// TIA Portal project "Project maybe not work 1.0" (V17) (continued)
REGION Network 7: step 20 Turns on intake and exhaust fans
   "Data_Block_Start_Seq".SeqStep[20] := "Data_Block_Start_Seq".StepNumber = 20;
   "Data_Block_Start_Seq".SeqConditions[20] := ("Data_Block_Start_Seq".StepNumber = 20) AND "FS-115.I" AND "FS-214-I" AND NOT "FS-114.I" AND NOT "FS-213.I" AND "HZ-413.I" AND NOT "PS-411.I" AND NOT "QE-116.I" AND "QE-316.I" AND NOT "Fire lock";
   "Data_Block_Start_Seq".SeqTimer[20].TON(IN := ("Data_Block_Start_Seq".StepNumber = 20) AND "Data_Block_Start_Seq".SeqConditions[20],
                           PT := T#50MS);
   IF "Data_Block_Start_Seq".SeqTimer[20].Q THEN
       "FC" := TRUE;
       "Data_Block_Start_Seq".StepNumber := 25;
   END_IF;
END_REGION

REGION Network 8: step 25 Checks that the fans have turned on
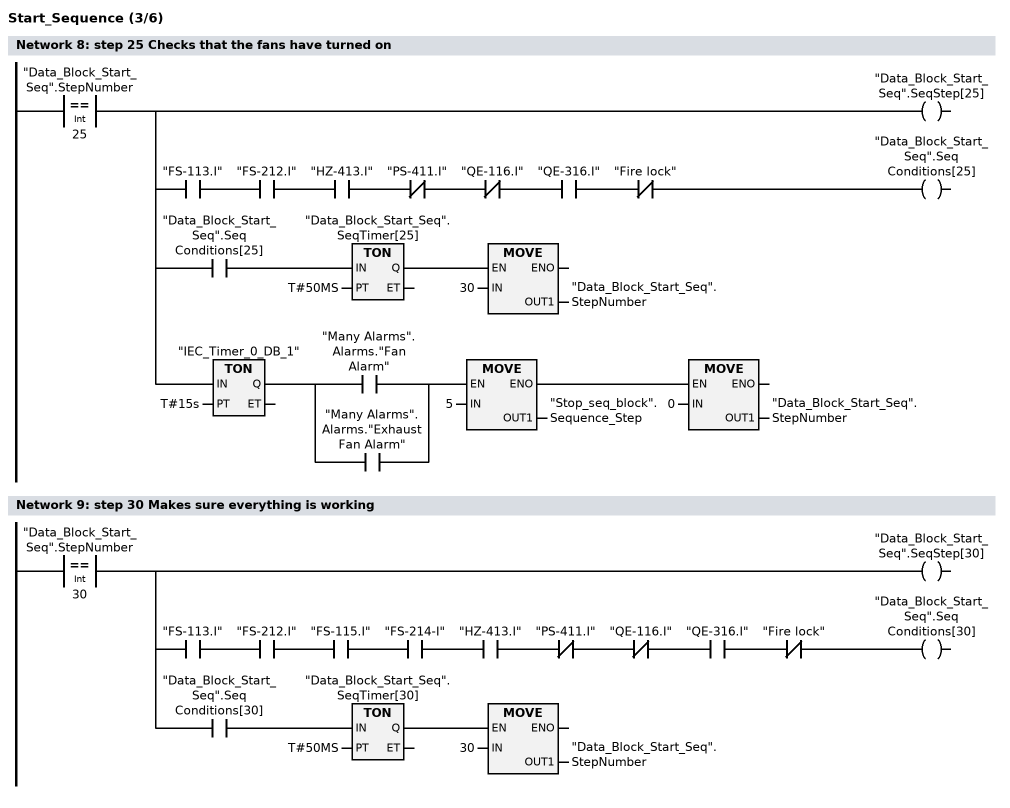
   "Data_Block_Start_Seq".SeqStep[25] := "Data_Block_Start_Seq".StepNumber = 25;
   "Data_Block_Start_Seq".SeqConditions[25] := ("Data_Block_Start_Seq".StepNumber = 25) AND "FS-113.I" AND "FS-212.I" AND "HZ-413.I" AND NOT "PS-411.I" AND NOT "QE-116.I" AND "QE-316.I" AND NOT "Fire lock";
   "Data_Block_Start_Seq".SeqTimer[25].TON(IN := ("Data_Block_Start_Seq".StepNumber = 25) AND "Data_Block_Start_Seq".SeqConditions[25],
                           PT := T#50MS);
   #_w1 := "Data_Block_Start_Seq".StepNumber = 25;
   IF "Data_Block_Start_Seq".SeqTimer[25].Q THEN "Data_Block_Start_Seq".StepNumber := 30; END_IF;
   "IEC_Timer_0_DB_1".TON(IN := #_w1, PT := T#15s);
   IF "IEC_Timer_0_DB_1".Q AND ("Many Alarms".Alarms."Fan Alarm" OR "Many Alarms".Alarms."Exhaust Fan Alarm") THEN
       "Stop_seq_block".Sequence_Step := 5;
       "Data_Block_Start_Seq".StepNumber := 0;
   END_IF;
END_REGION

REGION Network 9: step 30 Makes sure everything is working
   "Data_Block_Start_Seq".SeqStep[30] := "Data_Block_Start_Seq".StepNumber = 30;
   "Data_Block_Start_Seq".SeqConditions[30] := ("Data_Block_Start_Seq".StepNumber = 30) AND "FS-113.I" AND "FS-212.I" AND "FS-115.I" AND "FS-214-I" AND "HZ-413.I" AND NOT "PS-411.I" AND NOT "QE-116.I" AND "QE-316.I" AND NOT "Fire lock";
   "Data_Block_Start_Seq".SeqTimer[30].TON(IN := ("Data_Block_Start_Seq".StepNumber = 30) AND "Data_Block_Start_Seq".SeqConditions[30],
                           PT := T#50MS);
   IF "Data_Block_Start_Seq".SeqTimer[30].Q THEN "Data_Block_Start_Seq".StepNumber := 30; END_IF;
END_REGION

REGION Network 10: step 30 Makes sure everything is working
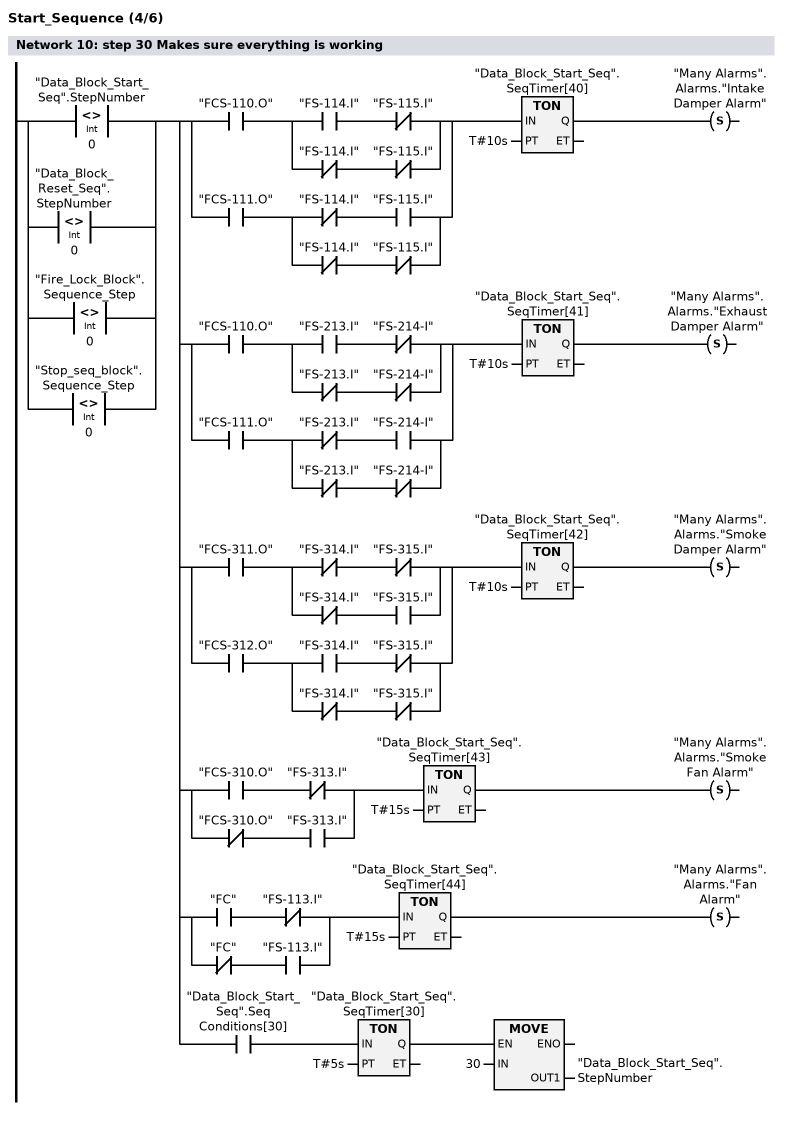
   #_w1 := ("Data_Block_Start_Seq".StepNumber <> 0) OR ("Data_Block_Reset_Seq".StepNumber <> 0) OR ("Fire_Lock_Block".Sequence_Step <> 0) OR ("Stop_seq_block".Sequence_Step <> 0);
   "Data_Block_Start_Seq".SeqTimer[40].TON(IN := #_w1 AND (("FCS-110.O" AND (("FS-114.I" AND NOT "FS-115.I") OR (NOT "FS-114.I" AND NOT "FS-115.I"))) OR ("FCS-111.O" AND ((NOT "FS-114.I" AND "FS-115.I") OR (NOT "FS-114.I" AND NOT "FS-115.I")))),
                           PT := T#10s);
   IF "Data_Block_Start_Seq".SeqTimer[40].Q THEN "Many Alarms".Alarms."Intake Damper Alarm" := TRUE; END_IF;
   "Data_Block_Start_Seq".SeqTimer[41].TON(IN := #_w1 AND (("FCS-110.O" AND (("FS-213.I" AND NOT "FS-214-I") OR (NOT "FS-213.I" AND NOT "FS-214-I"))) OR ("FCS-111.O" AND ((NOT "FS-213.I" AND "FS-214-I") OR (NOT "FS-213.I" AND NOT "FS-214-I")))),
                           PT := T#10s);
   IF "Data_Block_Start_Seq".SeqTimer[41].Q THEN "Many Alarms".Alarms."Exhaust Damper Alarm" := TRUE; END_IF;
   "Data_Block_Start_Seq".SeqTimer[42].TON(IN := #_w1 AND (("FCS-311.O" AND ((NOT "FS-314.I" AND NOT "FS-315.I") OR (NOT "FS-314.I" AND "FS-315.I"))) OR ("FCS-312.O" AND (("FS-314.I" AND NOT "FS-315.I") OR (NOT "FS-314.I" AND NOT "FS-315.I")))),
                           PT := T#10s);
   IF "Data_Block_Start_Seq".SeqTimer[42].Q THEN "Many Alarms".Alarms."Smoke Damper Alarm" := TRUE; END_IF;
   "Data_Block_Start_Seq".SeqTimer[43].TON(IN := #_w1 AND (("FCS-310.O" AND NOT "FS-313.I") OR (NOT "FCS-310.O" AND "FS-313.I")),
                           PT := T#15s);
   IF "Data_Block_Start_Seq".SeqTimer[43].Q THEN "Many Alarms".Alarms."Smoke Fan Alarm" := TRUE; END_IF;
   "Data_Block_Start_Seq".SeqTimer[44].TON(IN := #_w1 AND (("FC" AND NOT "FS-113.I") OR (NOT "FC" AND "FS-113.I")),
                           PT := T#15s);
   IF "Data_Block_Start_Seq".SeqTimer[44].Q THEN "Many Alarms".Alarms."Fan Alarm" := TRUE; END_IF;
   "Data_Block_Start_Seq".SeqTimer[30].TON(IN := #_w1 AND "Data_Block_Start_Seq".SeqConditions[30], PT := T#5s);
   IF "Data_Block_Start_Seq".SeqTimer[30].Q THEN "Data_Block_Start_Seq".StepNumber := 30; END_IF;
END_REGION

REGION Network 11: Stop and reset button function. after 3s puts on stop sequence if 10s passes reset function turns on
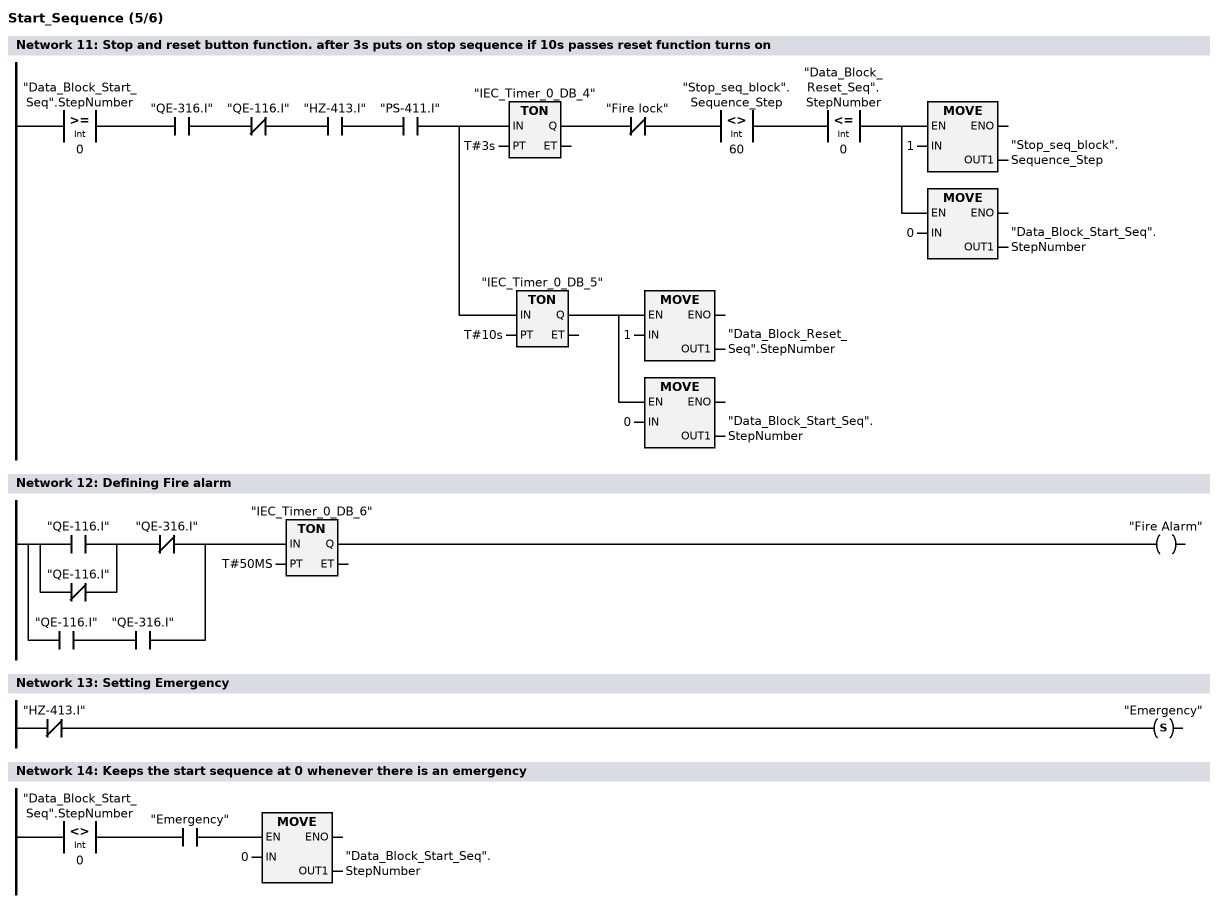
   #_w1 := ("Data_Block_Start_Seq".StepNumber >= 0) AND "QE-316.I" AND NOT "QE-116.I" AND "HZ-413.I" AND "PS-411.I";
   "IEC_Timer_0_DB_4".TON(IN := #_w1, PT := T#3s);
   #_w2 := "IEC_Timer_0_DB_4".Q AND NOT "Fire lock" AND ("Stop_seq_block".Sequence_Step <> 60) AND ("Data_Block_Reset_Seq".StepNumber <= 0);
   IF #_w2 THEN
       "Stop_seq_block".Sequence_Step := 1;
       "Data_Block_Start_Seq".StepNumber := 0;
   END_IF;
   "IEC_Timer_0_DB_5".TON(IN := #_w1, PT := T#10s);
   IF "IEC_Timer_0_DB_5".Q THEN
       "Data_Block_Reset_Seq".StepNumber := 1;
       "Data_Block_Start_Seq".StepNumber := 0;
   END_IF;
END_REGION

REGION Network 12: Defining Fire alarm
   "IEC_Timer_0_DB_6".TON(IN := (("QE-116.I" OR NOT "QE-116.I") AND NOT "QE-316.I") OR ("QE-116.I" AND "QE-316.I"),
                          PT := T#50MS);
   "Fire Alarm" := "IEC_Timer_0_DB_6".Q;
END_REGION

REGION Network 13: Setting Emergency
   RUNG wire#powerrail
      I_Contact( "HZ-413.I" )
      S_Coil( "Emergency" )
   END_RUNG
   // the same network as SCL:
   IF NOT "HZ-413.I" THEN "Emergency" := TRUE; END_IF;
END_REGION

REGION Network 14: Keeps the start sequence at 0 whenever there is an emergency
   RUNG wire#powerrail
      { S7_Templates := "SrcType := Int" } NE_Contact(in1 := "Data_Block_Start_Seq".StepNumber, in2 := 0)
      Contact( "Emergency" )
      Move(in := 0, out1 => "Data_Block_Start_Seq".StepNumber)
   END_RUNG
   // the same network as SCL:
   IF ("Data_Block_Start_Seq".StepNumber <> 0) AND "Emergency" THEN
       "Data_Block_Start_Seq".StepNumber := 0;
   END_IF;
END_REGION

REGION Network 15: Defining Alarm
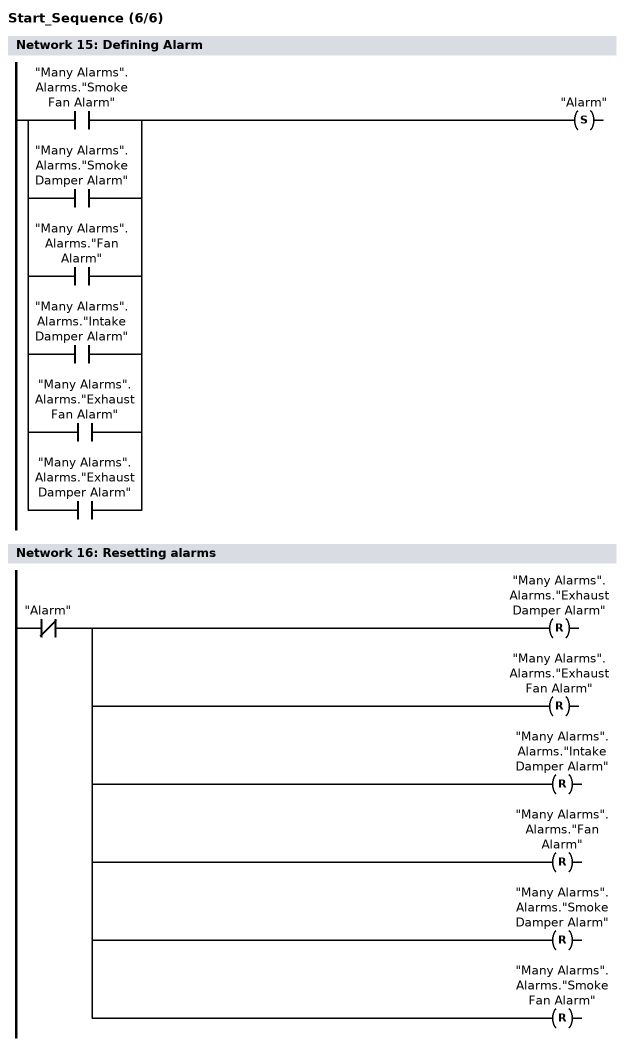
   RUNG wire#powerrail
      Contact( "Many Alarms".Alarms."Smoke Fan Alarm" )
      wire#w1
      S_Coil( "Alarm" )
   END_RUNG
   RUNG wire#powerrail
      Contact( "Many Alarms".Alarms."Smoke Damper Alarm" )
   END_RUNG wire#w1
   RUNG wire#powerrail
      Contact( "Many Alarms".Alarms."Fan Alarm" )
   END_RUNG wire#w1
   RUNG wire#powerrail
      Contact( "Many Alarms".Alarms."Intake Damper Alarm" )
   END_RUNG wire#w1
   RUNG wire#powerrail
      Contact( "Many Alarms".Alarms."Exhaust Fan Alarm" )
   END_RUNG wire#w1
   RUNG wire#powerrail
      Contact( "Many Alarms".Alarms."Exhaust Damper Alarm" )
   END_RUNG wire#w1
   // the same network as SCL:
   IF "Many Alarms".Alarms."Smoke Fan Alarm" OR "Many Alarms".Alarms."Smoke Damper Alarm" OR "Many Alarms".Alarms."Fan Alarm" OR "Many Alarms".Alarms."Intake Damper Alarm" OR "Many Alarms".Alarms."Exhaust Fan Alarm" OR "Many Alarms".Alarms."Exhaust Damper Alarm" THEN
       "Alarm" := TRUE;
   END_IF;
END_REGION

REGION Network 16: Resetting alarms
   RUNG wire#powerrail
      I_Contact( "Alarm" )
      wire#w1
      R_Coil( "Many Alarms".Alarms."Exhaust Damper Alarm" )
   END_RUNG
   RUNG wire#w1
      R_Coil( "Many Alarms".Alarms."Exhaust Fan Alarm" )
   END_RUNG
   RUNG wire#w1
      R_Coil( "Many Alarms".Alarms."Intake Damper Alarm" )
   END_RUNG
   RUNG wire#w1
      R_Coil( "Many Alarms".Alarms."Fan Alarm" )
   END_RUNG
   RUNG wire#w1
      R_Coil( "Many Alarms".Alarms."Smoke Damper Alarm" )
   END_RUNG
   RUNG wire#w1
      R_Coil( "Many Alarms".Alarms."Smoke Fan Alarm" )
   END_RUNG
   // the same network as SCL:
   IF NOT "Alarm" THEN
       "Many Alarms".Alarms."Exhaust Damper Alarm" := FALSE;
       "Many Alarms".Alarms."Exhaust Fan Alarm" := FALSE;
       "Many Alarms".Alarms."Intake Damper Alarm" := FALSE;
       "Many Alarms".Alarms."Fan Alarm" := FALSE;
       "Many Alarms".Alarms."Smoke Damper Alarm" := FALSE;
       "Many Alarms".Alarms."Smoke Fan Alarm" := FALSE;
   END_IF;
END_REGION
END_FUNCTION

ORGANIZATION_BLOCK "Main"   // OB1, LAD, ProgramCycle
TITLE = "Main Program Sweep (Cycle)"
{ S7_Optimized_Access := 'TRUE' }
VERSION : 0.1
   VAR_INPUT
      Initial_Call : Bool;   // Initial call of this OB
      Remanence : Bool;   // =True, if remanent data are available
   END_VAR
   VAR_TEMP
      "QE.200i-norm" : Real;
   END_VAR
   VAR_TEMP   // added for the SCL form of the ladder/FBD networks
      _w1 : Bool;
      _w2 : Bool;
      _w3 : Bool;
   END_VAR
BEGIN

REGION Network 1
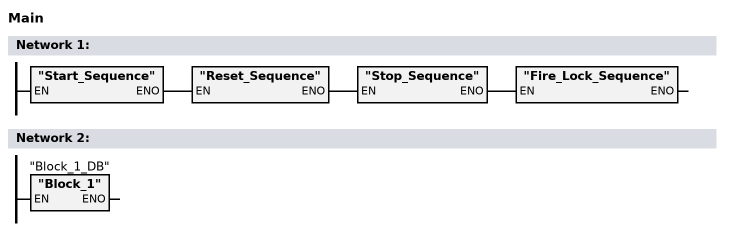
   RUNG wire#powerrail
      "Start_Sequence"()
      "Reset_Sequence"()
      "Stop_Sequence"()
      "Fire_Lock_Sequence"()
   END_RUNG
   // the same network as SCL:
   "Start_Sequence"(ENO => #_w1);
   "Reset_Sequence"(EN := #_w1, ENO => #_w2);
   "Stop_Sequence"(EN := #_w2, ENO => #_w3);
   IF #_w3 THEN "Fire_Lock_Sequence"(); END_IF;
END_REGION

REGION Network 2
   RUNG wire#powerrail
      "Block_1_DB"()
   END_RUNG
   // the same network as SCL:
   "Block_1_DB"();   // "Block_1"
END_REGION
END_ORGANIZATION_BLOCK

ORGANIZATION_BLOCK "Cyclic interrupt"   // OB30, LAD, CyclicInterrupt
{ S7_Optimized_Access := 'TRUE' }
VERSION : 0.1
   VAR_INPUT
      Initial_Call : Bool;   // Initial call of this OB
      Event_Count : Int;   // Events discarded
   END_VAR
   VAR_TEMP
      QE_Temp : Real;
      "TE temp" : Real;
      "TFC-Output temp" : Real;
   END_VAR
BEGIN

REGION Network 1
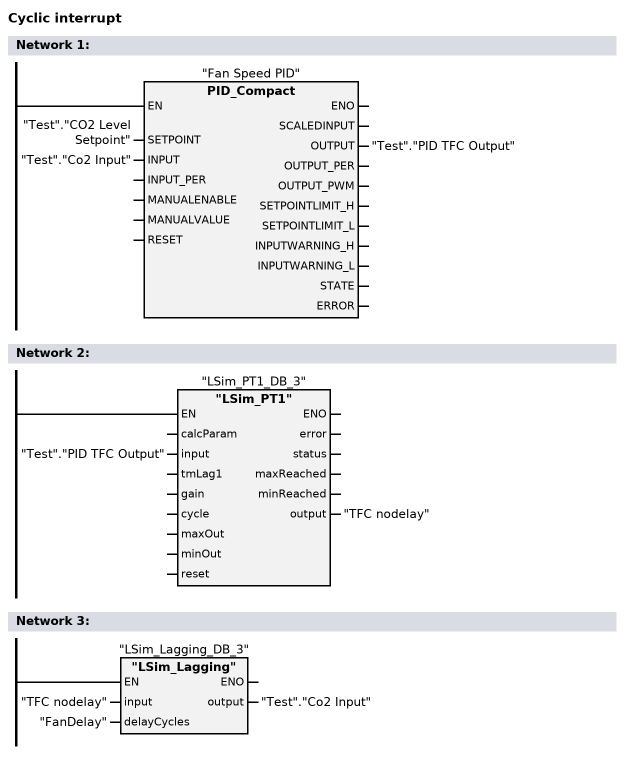
   "Fan Speed PID"(Setpoint := "Test"."CO2 Level Setpoint",   // PID_Compact
                   Input := "Test"."Co2 Input",
                   Output => "Test"."PID TFC Output");
END_REGION

REGION Network 2
   RUNG wire#powerrail
      "LSim_PT1_DB_3"(calcParam :=, input := "Test"."PID TFC Output", tmLag1 :=, gain :=, cycle :=, maxOut :=, minOut :=, reset :=, error =>, status =>, maxReached =>, minReached =>, output => "TFC nodelay")
   END_RUNG
   // the same network as SCL:
   "LSim_PT1_DB_3"(input := "Test"."PID TFC Output", output => "TFC nodelay");   // "LSim_PT1"
END_REGION

REGION Network 3
   RUNG wire#powerrail
      "LSim_Lagging_DB_3"(input := "TFC nodelay", delayCycles := "FanDelay", output => "Test"."Co2 Input")
   END_RUNG
   // the same network as SCL:
   "LSim_Lagging_DB_3"(input := "TFC nodelay", delayCycles := "FanDelay", output => "Test"."Co2 Input");   // "LSim_Lagging"
END_REGION
END_ORGANIZATION_BLOCK

ORGANIZATION_BLOCK "Cyclic interrupt_1"   // OB31, LAD, CyclicInterrupt
{ S7_Optimized_Access := 'TRUE' }
VERSION : 0.1
   VAR_INPUT
      Initial_Call : Bool;   // Initial call of this OB
      Event_Count : Int;   // Events discarded
   END_VAR
BEGIN

REGION Network 1
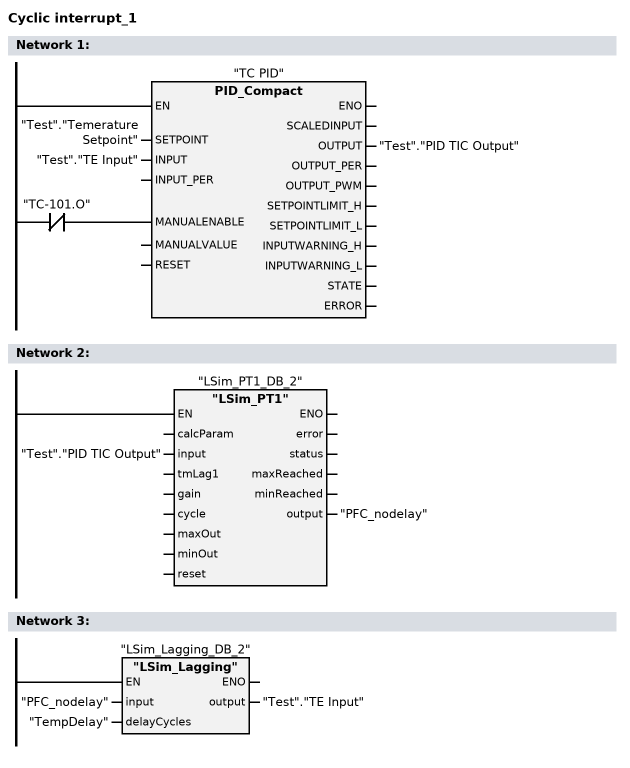
   "TC PID"(Setpoint := "Test"."Temerature Setpoint",   // PID_Compact
            Input := "Test"."TE Input",
            ManualEnable := NOT "TC-101.O",
            Output => "Test"."PID TIC Output");
END_REGION

REGION Network 2
   RUNG wire#powerrail
      "LSim_PT1_DB_2"(calcParam :=, input := "Test"."PID TIC Output", tmLag1 :=, gain :=, cycle :=, maxOut :=, minOut :=, reset :=, error =>, status =>, maxReached =>, minReached =>, output => "PFC_nodelay")
   END_RUNG
   // the same network as SCL:
   "LSim_PT1_DB_2"(input := "Test"."PID TIC Output", output => "PFC_nodelay");   // "LSim_PT1"
END_REGION

REGION Network 3
   RUNG wire#powerrail
      "LSim_Lagging_DB_2"(input := "PFC_nodelay", delayCycles := "TempDelay", output => "Test"."TE Input")
   END_RUNG
   // the same network as SCL:
   "LSim_Lagging_DB_2"(input := "PFC_nodelay", delayCycles := "TempDelay", output => "Test"."TE Input");   // "LSim_Lagging"
END_REGION
END_ORGANIZATION_BLOCK

(* ===== HMI "HMI_RT_1" =====
system functions are stored by id; their names below are inferred from use
connection "HMI_Connection_1": ETHERNET, S7_1200_OMS
connection "HMI_Connection_2": ETHERNET, S7_1200_OMS

HMI tags "Default tag table"
   "Tag_ScreenNumber" : UInt, internal
   "Fire lock" : Bool = PLC "Fire lock" AT %M36.2, 1 s
   "Emergency" : Bool = PLC Emergency AT %M36.4, 1 s
   "Intake Fan" : Bool = PLC "FS-113.I" AT %I6.1, 1 s
   "Exhaust Fan" : Bool = PLC "FS-212.I" AT %I6.4, 1 s
   "Intake Damper Closing" : Bool = PLC "FCS-111.O" AT %Q0.2, 1 s
   "Intake Damper Opening" : Bool = PLC "FCS-110.O" AT %Q0.1, 1 s
   "Intake Damper Closed" : Bool = PLC "FS-114.I" AT %I7.5, 1 s
   "Intake Damper Open" : Bool = PLC "FS-115.I" AT %I7.1, 1 s
   "Exhaust Damper Closing" : Bool = PLC "FCS-211.O" AT %Q0.4, 1 s
   "Exhaust Damper Closed" : Bool = PLC "FS-213.I" AT %I7.4, 1 s
   "Exhaust Damper Opening" : Bool = PLC "FCS-210O" AT %Q0.3, 1 s
   "Exhaust Damper Open" : Bool = PLC "FS-214-I" AT %I7.0, 1 s
   "Smoke Damper Opening" : Bool = PLC "FCS-311.O" AT %Q0.6, 1 s
   "Smoke Damper Open" : Bool = PLC "FS-314.I" AT %I7.2, 1 s
   "Smoke Damper Closing" : Bool = PLC "FCS-312.O" AT %Q0.7, 1 s
   "Smoke Damper Closed" : Bool = PLC "FS-315.I" AT %I7.6, 1 s
   "Smoke Fan Control" : Bool = PLC "FCS-310.O" AT %Q0.5, 1 s
   "Start Button" : Bool = PLC "PS-410.I" AT %I6.0, 1 s
   "Stop/Reset Button" : Bool = PLC "PS-411.I" AT %I6.3, 1 s
   "Emergency Button" : Bool = PLC "HZ-413.I" AT %I6.5, 1 s
   "Start Seq" : Int = PLC Data_Block_Start_Seq.StepNumber AT %DB1.DBX0.0, 1 s
   "Stop Seq" : Int = PLC Stop_seq_block.Sequence_Step AT %DB1.DBX0.0, 1 s
   "Reset Seq" : Int = PLC Data_Block_Reset_Seq.StepNumber AT %DB1.DBX0.0, 1 s
   "Fire Lock Seq" : Int = PLC Fire_Lock_Block.Sequence_Step AT %M36.2, 1 s
   "Fire Inside" : Bool = PLC "QE-316.I" AT %I7.7, 1 s
   "Fire Outside" : Bool = PLC "QE-116.I" AT %I7.3, 1 s
   "Smoke Fan Status" : Bool = PLC "FS-313.I" AT %I6.2, 1 s
   "Intake Fan Control" : Bool = PLC FC AT %M20.0, 1 s
   "Speed Scale" : Int = PLC Test."CO2 Level Setpoint" AT %DB1.DBW0, 1 s
   "TFC-201sp" : Real = PLC "Co2 Setpoint" AT %MD200, 1 s
   "QE-200.i" : Int = PLC "QE-200.i" AT %MW64, 1 s
   "TFC-201.o" : Real = PLC "TFC-201.o" AT %MD80, 1 s
   "Temperature.sp" : Int = PLC "Temperature.sp" AT %MW222, 1 s
   "TE-100.i" : Int = PLC "TE-100.i" AT %MW66, 1 s
   "TempratureSp" : Int = PLC "Temperature.sp" AT %MW222, 1 s
   "PFC-202.o" : Real = PLC "PFC-202.o" AT %MD84, 1 s
   "Test_PID_Data_Output" : Real = PLC Test."PID TFC Output", 1 s
   "Fan Speed PID_Output" : Real = PLC "Fan Speed PID".Output, 1 s
   "Fan Speed PID_Input" : Real = PLC "Fan Speed PID".Input, 1 s
   "Data_Block_Start_Seq_SeqStep{5}" : Bool = PLC Data_Block_Start_Seq.SeqStep[5], 1 s
   "Test_Temerature Setpoint" : Int = PLC Test."Temerature Setpoint", 1 s
   "TC PID_Input" : Real = PLC "TC PID".Input, 1 s
   "Fan Speed PID_State" : Int = PLC "Fan Speed PID".State, 1 s
   "TC PID_State" : Int = PLC "TC PID".State, 1 s

HMI tags "Alarms"
   "Alarms" : Int AT %DB4.DBW0, 1 s

discrete alarms
   1: 'Wha', class Warnings, trigger "Alarms" bit 0
   2: 'Wha', class Warnings, trigger "Alarms" bit 1
   3: 'Wha', class Warnings, trigger "Alarms" bit 2
   4: 'Wha', class Warnings, trigger "Alarms" bit 3
   5: 'Wha', class Warnings, trigger "Alarms" bit 4
   6: 'Wha', class Warnings, trigger "Alarms" bit 5
   7: 'Wha', class Warnings, trigger "Alarms" bit 6
   8: 'Wha', class Warnings, trigger "Alarms" bit 7
   9: 'Intake Damper Control Time Exceeded', class Errors, trigger "Alarms" bit 8
   10: 'Intake Fan Control Time Exceeded', class Errors, trigger "Alarms" bit 9
   13: 't Dameper Control Time Exceeded', class Errors, trigger "Alarms" bit 10
   14: 'Exhaust Fan Control time Exceeded', class Errors, trigger "Alarms" bit 11
   15: 'Smoke Damper Control Time Exceeded', class Errors, trigger "Alarms" bit 12
   16: 'Smoke Fan Control Time Exceeded', class Errors, trigger "Alarms" bit 13

screen "Root screen" 1280x757, template "Template_1"
   on GenerateScreen: SetTag("Tag_ScreenNumber", 1)
   Circle "Circle_1" at 336,50 size 29x29
      Appearance <- "Fire lock"
   Circle "Circle_2" at 334,83 size 29x29
      Appearance <- "Emergency"
      Visibility <- "Emergency"
   Button "HmiScreenItemData_2" at 36,95 size 159x47; TextOff 'System screens'; PictureOff "Navigates to System screens for TP2200 Comfort V2 17.0.0.0"; PictureOn "Navigates to System screens for TP2200 Comfort V2 17.0.0.0"
      on Release: ActivateScreen("System screens", 0)
   Button "HmiScreenItemData" at 36,36 size 159x47; TextOff 'Screen0'; PictureOff "Navigates to Screen0 for TP2200 Comfort V2 17.0.0.0"; PictureOn "Navigates to Screen0 for TP2200 Comfort V2 17.0.0.0"
      on Release: ActivateScreen("Screen0", 0)
   Rectangle "Exhaust Damper Opening" at 833,244 size 54x23
      Appearance <- "Exhaust Damper Opening"
      Visibility <- "Exhaust Damper Opening"
   Rectangle "Intake Damper Opening" at 542,400 size 54x23
      Appearance <- "Intake Damper Opening"
      Visibility <- "Intake Damper Opening"
   Rectangle "Intake Damper Closing" at 542,400 size 54x23
      Appearance <- "Intake Damper Closing"
      Visibility <- "Intake Damper Closing"
   Rectangle "Exhaust Damper Closing" at 833,244 size 54x23
      Appearance <- "Exhaust Damper Closing"
      Visibility <- "Exhaust Damper Closing"
   Circle "Circle_3" at 334,83 size 29x29
      Appearance <- "Emergency Button"
      Visibility <- "Emergency Button"
   Rectangle "Smoke Damper Closing" at 833,149 size 54x23
      Appearance <- "Smoke Damper Closing"
      Visibility <- "Smoke Damper Closing"
   Rectangle "Smoke Damper Opening" at 833,149 size 54x23
      Appearance <- "Smoke Damper Opening"
      Visibility <- "Smoke Damper Opening"
   Button "Smoke Damper Closed Button_1" at 210,565 size 96x32; TextOff 'Closed'
      on Click: SetBit("Smoke Damper Closed")
      Visibility <- "Smoke Damper Closed"
   Button "Smoke Damper Open Button_1" at 210,610 size 96x32; TextOff 'Open'
      on Click: SetBit("Smoke Damper Open")
      Visibility <- "Smoke Damper Open"
   Button "Smoke Damper Not Closed Button_1" at 210,566 size 96x32; TextOff 'Not Closed'
      on Click: ResetBit("Smoke Damper Closed")
      Visibility <- "Smoke Damper Closed"
   Button "Smoke Damper Not Open Button_1" at 210,609 size 96x32; TextOff 'Not Open'
      on Click: ResetBit("Smoke Damper Open")
      Visibility <- "Smoke Damper Open"
   Button "Intake Damper Closed Button" at 7,565 size 96x32; TextOff 'Closed'
      on Click: SetBit("Intake Damper Closed")
      Visibility <- "Intake Damper Closed"
   Button "Intake Damper Open Button" at 7,610 size 96x32; TextOff 'Open'
      on Click: SetBit("Intake Damper Open")
      Visibility <- "Intake Damper Open"
   Button "Intake Damper Not Closed Button" at 8,565 size 96x32; TextOff 'Not Closed'
      on Click: ResetBit("Intake Damper Closed")
      Visibility <- "Intake Damper Closed"
   Button "Exhaust Damper Closed Button" at 108,565 size 96x32; TextOff 'Closed'
      on Click: SetBit("Exhaust Damper Closed")
      Visibility <- "Exhaust Damper Closed"
   Button "Intake Damper Not Open Button" at 7,608 size 96x32; TextOff 'Not Open'
      Visibility <- "Intake Damper Open"
      on Click: ResetBit("Intake Damper Open")
   Button "Exhaust Damper Open Button" at 108,610 size 96x32; TextOff 'Open'
      on Click: SetBit("Exhaust Damper Open")
      Visibility <- "Exhaust Damper Open"
   Button "Exhaust Damper Not Closed Button" at 108,565 size 96x32; TextOff 'Not Closed'
      on Click: ResetBit("Exhaust Damper Closed")
      Visibility <- "Exhaust Damper Closed"
   Button "Exhaust Damper Not Open Button" at 108,608 size 96x32; TextOff 'Not Open'
      on Click: ResetBit("Exhaust Damper Open")
      Visibility <- "Exhaust Damper Open"
   GraphicView "Graphic view_1" at 430,120 size 824x564; Picture "Graphic_10"
   Rectangle "Exhaust Fan" at 650,229 size 54x23
      Appearance <- "Intake Fan Control"
   Rectangle "Intake Fan" at 730,383 size 54x23
      Appearance <- "Intake Fan Control"
   Rectangle "Intake Damper Closed" at 542,400 size 54x23
      Appearance <- "Intake Damper Closed"
      Visibility <- "Intake Damper Closed"
   Rectangle "Intake Damper Open" at 542,400 size 54x23
      Appearance <- "Intake Damper Open"
      Visibility <- "Intake Damper Open"
   Rectangle "Exhaust Damper Open" at 833,244 size 54x23
      Appearance <- "Exhaust Damper Open"
      Visibility <- "Exhaust Damper Open"
   Rectangle "Exhaust Damper Closed" at 833,244 size 54x23
      Visibility <- "Exhaust Damper Closed"
      Appearance <- "Exhaust Damper Closed"
   Rectangle "Smoke Damper Open" at 833,149 size 54x23
      Appearance <- "Smoke Damper Open"
      Visibility <- "Smoke Damper Open"
   Rectangle "Smoke Damper Closed" at 833,149 size 54x23
      Visibility <- "Smoke Damper Closed"
      Appearance <- "Smoke Damper Closed"
   Button "Intake Fan Off" at 7,648 size 96x32; TextOff 'OFF'
      on Click: ResetBit("Intake Fan")
      Visibility <- "Intake Fan"
   Button "Intake Fan On" at 7,648 size 96x32; TextOff 'ON'
      on Click: SetBit("Intake Fan")
      Visibility <- "Intake Fan"
   Button "Exhaust Fan Off" at 108,648 size 96x32; TextOff 'OFF'
      on Click: ResetBit("Exhaust Fan")
      Visibility <- "Exhaust Fan"
   Button "Exhaust Fan on" at 108,648 size 96x32; TextOff 'ON'
      on Click: SetBit("Exhaust Fan")
      Visibility <- "Exhaust Fan"
   Button "Button_1" at 47,162 size 210x95; TextOff 'Start'
      on Press: SetBit("Start Button")
      on Release: ResetBit("Start Button")
      Appearance <- "Data_Block_Start_Seq_SeqStep{5}"
   Button "Button_2" at 47,272 size 210x45; TextOff 'Stop/Reset'
      on Press: SetBit("Stop/Reset Button")
      on Release: ResetBit("Stop/Reset Button")
   Button "Button_3" at 45,340 size 210x45; TextOff 'Release Emergency'
      on Click: SetBit("Emergency Button")
   Button "Button_4" at 45,387 size 210x45; TextOff 'Emergency'
      on Click: ResetBit("Emergency Button")
   Rectangle "Rectangle_1" at 416,67 size 50x45
      Appearance <- "Start Seq"
   Rectangle "Rectangle_2" at 479,65 size 50x45
      Appearance <- "Stop Seq"
   Rectangle "Rectangle_3" at 544,67 size 50x45
      Appearance <- "Reset Seq"
   Rectangle "Rectangle_4" at 607,65 size 50x45
      Appearance <- "Fire Lock Seq"
   Button "Button_5" at 35,480 size 96x32; TextOff 'Fire O'
      on Click: SetBit("Fire Outside")
      Visibility <- "Fire Outside"
   Button "Button_6" at 32,480 size 96x32; TextOff 'No Fire O'
      on Click: ResetBit("Fire Outside")
      Visibility <- "Fire Outside"
   Button "Button_7" at 177,480 size 96x32; TextOff 'Fire I'
      on Click: ResetBit("Fire Inside")
      Visibility <- "Fire Inside"
   Button "Button_8" at 178,480 size 96x32; TextOff 'No Fire I'
      on Click: SetBit("Fire Inside")
      Visibility <- "Fire Inside"
   Rectangle "Rectangle_5" at 35,443 size 95x24
      Appearance <- "Fire Outside"
   Rectangle "Rectangle_6" at 180,442 size 95x24
      Appearance <- "Fire Inside"
   Rectangle "Smoke Exhaust Fan_1" at 652,133 size 54x23
      Appearance <- "Smoke Fan Control"
   TextField "Text field_1" at 23,540 size 67x25; Text 'Intake'
   TextField "Text field_2" at 115,540 size 80x25; Text 'Exhaust'
   TextField "Text field_3" at 225,540 size 68x25; Text 'Smoke'
   Button "Smoke Fan Off" at 210,648 size 96x32; TextOff 'OFF'
      on Click: ResetBit("Smoke Fan Status")
      Visibility <- "Smoke Fan Status"
   Button "Smoke Fan On" at 210,648 size 96x32; TextOff 'ON'
      on Click: SetBit("Smoke Fan Status")
      Visibility <- "Smoke Fan Status"
   Button "Button_10" at 649,256 size 64x61; TextOff 'Text'; TextOn 'Exhaust Fan Speed'
      on Click: function_efd93a16("Fan Speed", 0, 0, -1, -1, 1)
   Button "Button_11" at 890,402 size 151x79; TextOff 'Text'; TextOn 'Pop-up screen_1'
      on Click: function_efd93a16("Pop-up screen_1", 0, 0, -1, -1, 1)
   Bar "Bar_1" at 1147,164 size 80x230; MinimumValue 0; MaximumValue 100
      ProcessValue <- "Fan Speed PID_Input"
   IOField "I/O field_1" at 1142,405 size 96x32; FormatPattern 999; Unit %
      ProcessValue <- "Speed Scale"
   TextField "Text field_4" at 1162,138 size 43x25; Text 'CO2'
   Button "Button_9" at 733,412 size 55x58; TextOn 'Exhaust Fan Speed'; TextOff 'Text'
      on Click: function_efd93a16("Fan Speed", 0, 0, -1, -1, 1)
   IOField "I/O field_2" at 1142,459 size 96x32; FormatPattern s99999
      ProcessValue <- "Fan Speed PID_State"
   IOField "I/O field_3" at 919,488 size 96x32; FormatPattern s99999
      ProcessValue <- "TC PID_State"

screen "Screen0" 1280x757, template "Template_1"
   on GenerateScreen: SetTag("Tag_ScreenNumber", 2)
   Button "Back" at 1,1 size 159x47; TextOff 'Back'
      on Release: ActivateScreen("Root screen", 0)
   AlarmView "Alarm view_1" at 4,48 size 1103x611

screen "System screens" 1280x757, template "Template_1"
   on GenerateScreen: SetTag("Tag_ScreenNumber", 3)
   Button "Back" at 1,1 size 159x47; TextOff 'Back'
      on Release: ActivateScreen("Root screen", 0)

PopupScreen "Fan Speed" 240x240
   Bar "Bar_1" at 0,92 size 240x72; MinimumValue 20; MaximumValue 100
      ProcessValue <- "Fan Speed PID_Output"

PopupScreen "Pop-up screen_1" 240x240
   Slider "Slider_1" at 0,108 size 239x68; Caption 'SIMATIC'
      ProcessValue <- "Test_Temerature Setpoint"
   Bar "Bar_1" at 0,34 size 239x65; MinimumValue 0; MaximumValue 50
      ProcessValue <- "TC PID_Input"

Template "Template_1" 1280x757
   Button "Exit" at 1200,679 size 78x59; TextOn 'Exit'; TextOff 'Exit'; PictureOn "ExitRuntime_TP1500_Comfort_V2_TR"; PictureOff "ExitRuntime_TP1500_Comfort_V2_TR"
      on Release: StopRuntime(0)
   Button "Template_Button" at 1120,679 size 78x59; TextOff 'Text'
   Button "Template_Button_1" at 1040,679 size 78x59; TextOff 'Text'
   Button "Template_Button_2" at 960,679 size 78x59; TextOff 'Text'
   Button "Template_Button_3" at 880,679 size 78x59; TextOff 'Text'
   Button "Template_Button_4" at 800,679 size 78x59; TextOff 'Text'
   Button "Template_Button_5" at 720,679 size 78x59; TextOff 'Text'
   Button "Template_Button_6" at 640,679 size 78x59; TextOff 'Text'
   Button "Template_Button_7" at 561,679 size 78x59; TextOff 'Text'
   Button "Template_Button_8" at 481,679 size 78x59; TextOff 'Text'
   Button "Template_Button_9" at 401,679 size 78x59; TextOff 'Text'
   Button "Template_Button_10" at 321,679 size 78x59; TextOff 'Text'
   Button "Template_Button_11" at 241,679 size 78x59; TextOff 'Text'
   Button "Template_Button_12" at 161,679 size 78x59; TextOff 'Text'
   Button "Alarms" at 81,679 size 78x59; TextOn 'Alarms'; TextOff 'Alarms'; PictureOn "AlarmDisplay_TP1500_Comfort_V2_TR"; PictureOff "AlarmDisplay_TP1500_Comfort_V2_TR"
      on Release: function_ef3f5d25("Alarm window_Unacknowledged", -1)
   Button "Start screen" at 1,679 size 78x59; TextOn 'Start screen'; TextOff 'Start screen'; PictureOn "NavigateHome_TP1500_Comfort_V2_TR"; PictureOff "NavigateHome_TP1500_Comfort_V2_TR"
      on Release: ActivateScreen("Root screen", 0)
*)